VERSION : 0.1
   VAR_TEMP   // added for the SCL form of the ladder/FBD networks
      _w1 : Bool;
      _s5time1 : S5Time;
   END_VAR
BEGIN

REGION Network 1: Aviso 1 - Falla Conexión con sensor de Temperatura torres de Cavaleto
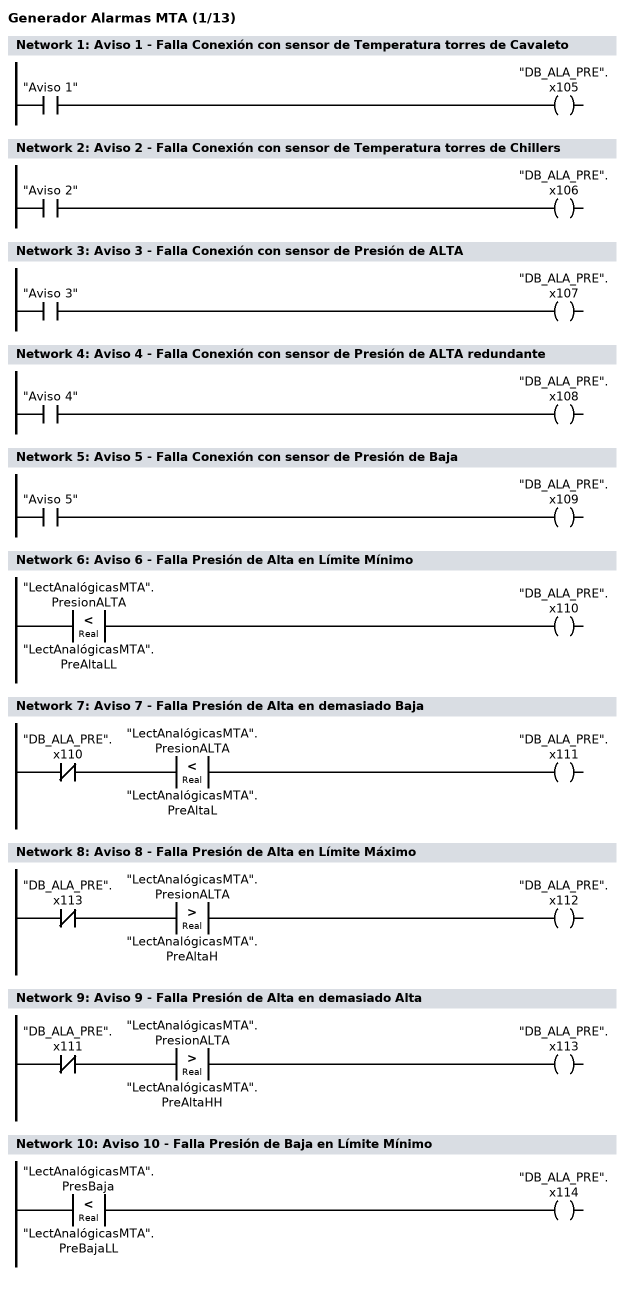
   RUNG wire#powerrail
      Contact( "Aviso 1" )
      Coil( "DB_ALA_PRE".x105 )
   END_RUNG
   // the same network as SCL:
   "DB_ALA_PRE".x105 := "Aviso 1";
END_REGION

REGION Network 2: Aviso 2 - Falla Conexión con sensor de Temperatura torres de Chillers
   RUNG wire#powerrail
      Contact( "Aviso 2" )
      Coil( "DB_ALA_PRE".x106 )
   END_RUNG
   // the same network as SCL:
   "DB_ALA_PRE".x106 := "Aviso 2";
END_REGION

REGION Network 3: Aviso 3 - Falla Conexión con sensor de Presión de ALTA
   RUNG wire#powerrail
      Contact( "Aviso 3" )
      Coil( "DB_ALA_PRE".x107 )
   END_RUNG
   // the same network as SCL:
   "DB_ALA_PRE".x107 := "Aviso 3";
END_REGION

REGION Network 4: Aviso 4 - Falla Conexión con sensor de Presión de ALTA redundante
   RUNG wire#powerrail
      Contact( "Aviso 4" )
      Coil( "DB_ALA_PRE".x108 )
   END_RUNG
   // the same network as SCL:
   "DB_ALA_PRE".x108 := "Aviso 4";
END_REGION

REGION Network 5: Aviso 5 - Falla Conexión con sensor de Presión de Baja
   RUNG wire#powerrail
      Contact( "Aviso 5" )
      Coil( "DB_ALA_PRE".x109 )
   END_RUNG
   // the same network as SCL:
   "DB_ALA_PRE".x109 := "Aviso 5";
END_REGION

REGION Network 6: Aviso 6 - Falla Presión de Alta en Límite Mínimo
   RUNG wire#powerrail
      { S7_Templates := "SrcType := Real" } LT_Contact(in1 := "LectAnalógicasMTA".PresionALTA, in2 := "LectAnalógicasMTA".PreAltaLL)
      Coil( "DB_ALA_PRE".x110 )
   END_RUNG
   // the same network as SCL:
   "DB_ALA_PRE".x110 := "LectAnalógicasMTA".PresionALTA < "LectAnalógicasMTA".PreAltaLL;
END_REGION

REGION Network 7: Aviso 7 - Falla Presión de Alta en demasiado Baja
   RUNG wire#powerrail
      I_Contact( "DB_ALA_PRE".x110 )
      { S7_Templates := "SrcType := Real" } LT_Contact(in1 := "LectAnalógicasMTA".PresionALTA, in2 := "LectAnalógicasMTA".PreAltaL)
      Coil( "DB_ALA_PRE".x111 )
   END_RUNG
   // the same network as SCL:
   "DB_ALA_PRE".x111 := NOT "DB_ALA_PRE".x110 AND ("LectAnalógicasMTA".PresionALTA < "LectAnalógicasMTA".PreAltaL);
END_REGION

REGION Network 8: Aviso 8 - Falla Presión de Alta en Límite Máximo
   RUNG wire#powerrail
      I_Contact( "DB_ALA_PRE".x113 )
      { S7_Templates := "SrcType := Real" } GT_Contact(in1 := "LectAnalógicasMTA".PresionALTA, in2 := "LectAnalógicasMTA".PreAltaH)
      Coil( "DB_ALA_PRE".x112 )
   END_RUNG
   // the same network as SCL:
   "DB_ALA_PRE".x112 := NOT "DB_ALA_PRE".x113 AND ("LectAnalógicasMTA".PresionALTA > "LectAnalógicasMTA".PreAltaH);
END_REGION

REGION Network 9: Aviso 9 - Falla Presión de Alta en demasiado Alta
   RUNG wire#powerrail
      I_Contact( "DB_ALA_PRE".x111 )
      { S7_Templates := "SrcType := Real" } GT_Contact(in1 := "LectAnalógicasMTA".PresionALTA, in2 := "LectAnalógicasMTA".PreAltaHH)
      Coil( "DB_ALA_PRE".x113 )
   END_RUNG
   // the same network as SCL:
   "DB_ALA_PRE".x113 := NOT "DB_ALA_PRE".x111 AND ("LectAnalógicasMTA".PresionALTA > "LectAnalógicasMTA".PreAltaHH);
END_REGION

REGION Network 10: Aviso 10 - Falla Presión de Baja en Límite Mínimo
   RUNG wire#powerrail
      { S7_Templates := "SrcType := Real" } LT_Contact(in1 := "LectAnalógicasMTA".PresBaja, in2 := "LectAnalógicasMTA".PreBajaLL)
      Coil( "DB_ALA_PRE".x114 )
   END_RUNG
   // the same network as SCL:
   "DB_ALA_PRE".x114 := "LectAnalógicasMTA".PresBaja < "LectAnalógicasMTA".PreBajaLL;
END_REGION

REGION Network 11: Aviso 11 - Falla Presión de Baja en demasiado Baja
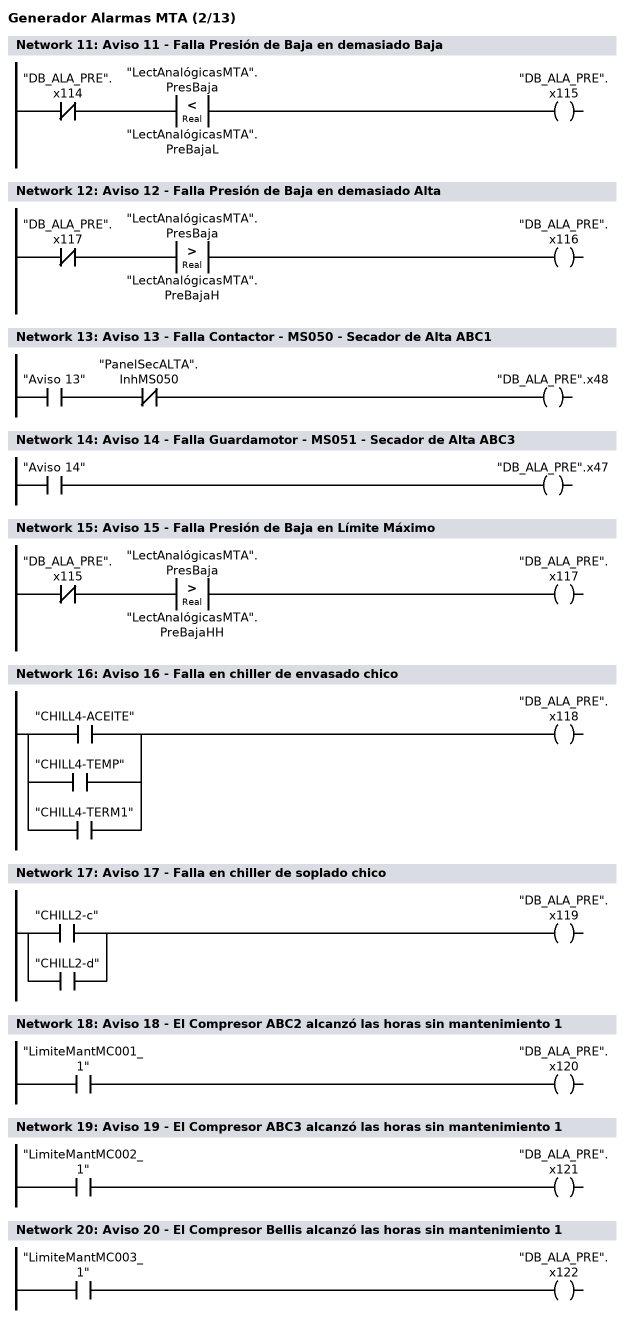
   RUNG wire#powerrail
      I_Contact( "DB_ALA_PRE".x114 )
      { S7_Templates := "SrcType := Real" } LT_Contact(in1 := "LectAnalógicasMTA".PresBaja, in2 := "LectAnalógicasMTA".PreBajaL)
      Coil( "DB_ALA_PRE".x115 )
   END_RUNG
   // the same network as SCL:
   "DB_ALA_PRE".x115 := NOT "DB_ALA_PRE".x114 AND ("LectAnalógicasMTA".PresBaja < "LectAnalógicasMTA".PreBajaL);
END_REGION

REGION Network 12: Aviso 12 - Falla Presión de Baja en demasiado Alta
   RUNG wire#powerrail
      I_Contact( "DB_ALA_PRE".x117 )
      { S7_Templates := "SrcType := Real" } GT_Contact(in1 := "LectAnalógicasMTA".PresBaja, in2 := "LectAnalógicasMTA".PreBajaH)
      Coil( "DB_ALA_PRE".x116 )
   END_RUNG
   // the same network as SCL:
   "DB_ALA_PRE".x116 := NOT "DB_ALA_PRE".x117 AND ("LectAnalógicasMTA".PresBaja > "LectAnalógicasMTA".PreBajaH);
END_REGION

REGION Network 13: Aviso 13 - Falla Contactor - MS050 - Secador de Alta ABC1
   RUNG wire#powerrail
      Contact( "Aviso 13" )
      I_Contact( "PanelSecALTA".InhMS050 )
      Coil( "DB_ALA_PRE".x48 )
   END_RUNG
   // the same network as SCL:
   "DB_ALA_PRE".x48 := "Aviso 13" AND NOT "PanelSecALTA".InhMS050;
END_REGION

REGION Network 14: Aviso 14 - Falla Guardamotor - MS051 - Secador de Alta ABC3
   RUNG wire#powerrail
      Contact( "Aviso 14" )
      Coil( "DB_ALA_PRE".x47 )
   END_RUNG
   // the same network as SCL:
   "DB_ALA_PRE".x47 := "Aviso 14";
END_REGION

REGION Network 15: Aviso 15 - Falla Presión de Baja en Límite Máximo
   RUNG wire#powerrail
      I_Contact( "DB_ALA_PRE".x115 )
      { S7_Templates := "SrcType := Real" } GT_Contact(in1 := "LectAnalógicasMTA".PresBaja, in2 := "LectAnalógicasMTA".PreBajaHH)
      Coil( "DB_ALA_PRE".x117 )
   END_RUNG
   // the same network as SCL:
   "DB_ALA_PRE".x117 := NOT "DB_ALA_PRE".x115 AND ("LectAnalógicasMTA".PresBaja > "LectAnalógicasMTA".PreBajaHH);
END_REGION

REGION Network 16: Aviso 16 - Falla en chiller de envasado chico
   RUNG wire#powerrail
      Contact( "CHILL4-ACEITE" )
      wire#w1
      Coil( "DB_ALA_PRE".x118 )
   END_RUNG
   RUNG wire#powerrail
      Contact( "CHILL4-TEMP" )
   END_RUNG wire#w1
   RUNG wire#powerrail
      Contact( "CHILL4-TERM1" )
   END_RUNG wire#w1
   // the same network as SCL:
   "DB_ALA_PRE".x118 := "CHILL4-ACEITE" OR "CHILL4-TEMP" OR "CHILL4-TERM1";
END_REGION

REGION Network 17: Aviso 17 - Falla en chiller de soplado chico
   RUNG wire#powerrail
      Contact( "CHILL2-c" )
      wire#w1
      Coil( "DB_ALA_PRE".x119 )
   END_RUNG
   RUNG wire#powerrail
      Contact( "CHILL2-d" )
   END_RUNG wire#w1
   // the same network as SCL:
   "DB_ALA_PRE".x119 := "CHILL2-c" OR "CHILL2-d";
END_REGION

REGION Network 18: Aviso 18 - El Compresor ABC2 alcanzó las horas sin mantenimiento 1
   RUNG wire#powerrail
      Contact( "LimiteMantMC001_1" )
      Coil( "DB_ALA_PRE".x120 )
   END_RUNG
   // the same network as SCL:
   "DB_ALA_PRE".x120 := "LimiteMantMC001_1";
END_REGION

REGION Network 19: Aviso 19 - El Compresor ABC3 alcanzó las horas sin mantenimiento 1
   RUNG wire#powerrail
      Contact( "LimiteMantMC002_1" )
      Coil( "DB_ALA_PRE".x121 )
   END_RUNG
   // the same network as SCL:
   "DB_ALA_PRE".x121 := "LimiteMantMC002_1";
END_REGION

REGION Network 20: Aviso 20 - El Compresor Bellis alcanzó las horas sin mantenimiento 1
   RUNG wire#powerrail
      Contact( "LimiteMantMC003_1" )
      Coil( "DB_ALA_PRE".x122 )
   END_RUNG
   // the same network as SCL:
   "DB_ALA_PRE".x122 := "LimiteMantMC003_1";
END_REGION

REGION Network 21: Aviso 21 - El Compresor ABC4 alcanzó las horas sin mantenimiento 1
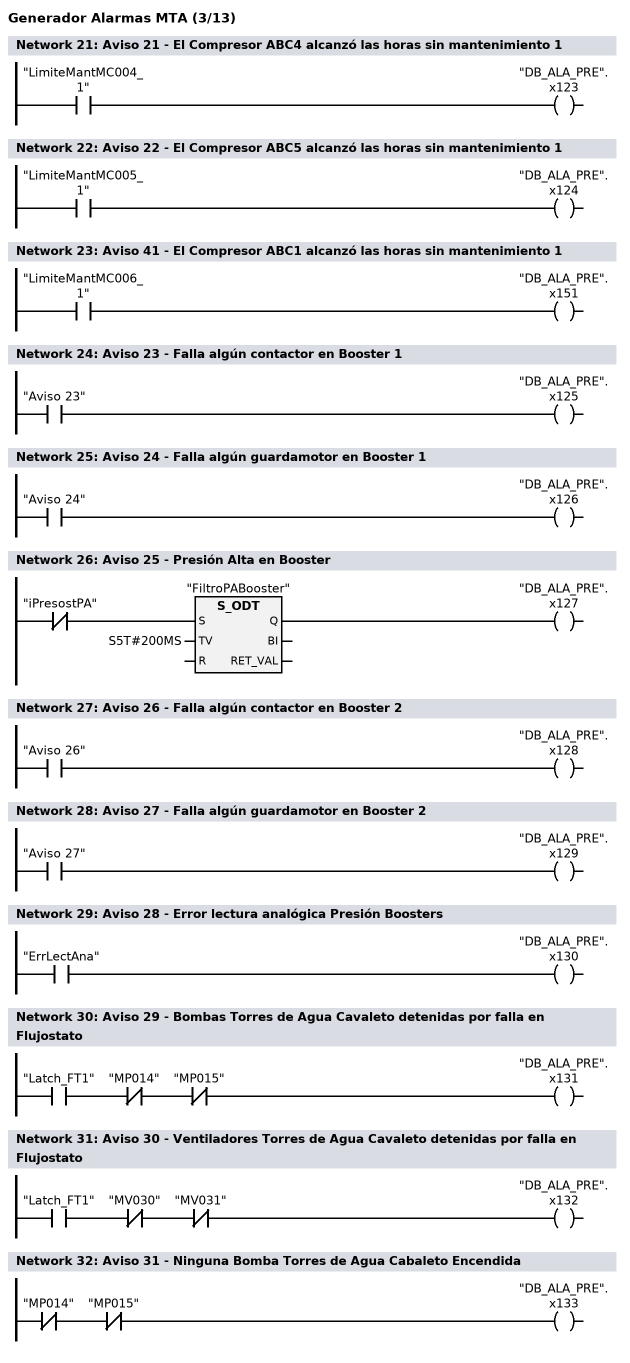
   RUNG wire#powerrail
      Contact( "LimiteMantMC004_1" )
      Coil( "DB_ALA_PRE".x123 )
   END_RUNG
   // the same network as SCL:
   "DB_ALA_PRE".x123 := "LimiteMantMC004_1";
END_REGION

REGION Network 22: Aviso 22 - El Compresor ABC5 alcanzó las horas sin mantenimiento 1
   RUNG wire#powerrail
      Contact( "LimiteMantMC005_1" )
      Coil( "DB_ALA_PRE".x124 )
   END_RUNG
   // the same network as SCL:
   "DB_ALA_PRE".x124 := "LimiteMantMC005_1";
END_REGION

REGION Network 23: Aviso 41 - El Compresor ABC1 alcanzó las horas sin mantenimiento 1
   RUNG wire#powerrail
      Contact( "LimiteMantMC006_1" )
      Coil( "DB_ALA_PRE".x151 )
   END_RUNG
   // the same network as SCL:
   "DB_ALA_PRE".x151 := "LimiteMantMC006_1";
END_REGION

REGION Network 24: Aviso 23 - Falla algún contactor en Booster 1
   RUNG wire#powerrail
      Contact( "Aviso 23" )
      Coil( "DB_ALA_PRE".x125 )
   END_RUNG
   // the same network as SCL:
   "DB_ALA_PRE".x125 := "Aviso 23";
END_REGION

REGION Network 25: Aviso 24 - Falla algún guardamotor en Booster 1
   RUNG wire#powerrail
      Contact( "Aviso 24" )
      Coil( "DB_ALA_PRE".x126 )
   END_RUNG
   // the same network as SCL:
   "DB_ALA_PRE".x126 := "Aviso 24";
END_REGION

REGION Network 26: Aviso 25 - Presión Alta en Booster
   RUNG wire#powerrail
      I_Contact( "iPresostPA" )
      S_ODT(T_NO := "FiltroPABooster", TV := S5T#200MS, R :=, BI =>, RET_VAL =>)
      Coil( "DB_ALA_PRE".x127 )
   END_RUNG
   // the same network as SCL:
   #_s5time1 := S_ODT(T_NO := "FiltroPABooster", S := NOT "iPresostPA", TV := S5T#200MS, Q => #_w1);
   "DB_ALA_PRE".x127 := #_w1;
END_REGION

REGION Network 27: Aviso 26 - Falla algún contactor en Booster 2
   RUNG wire#powerrail
      Contact( "Aviso 26" )
      Coil( "DB_ALA_PRE".x128 )
   END_RUNG
   // the same network as SCL:
   "DB_ALA_PRE".x128 := "Aviso 26";
END_REGION

REGION Network 28: Aviso 27 - Falla algún guardamotor en Booster 2
   RUNG wire#powerrail
      Contact( "Aviso 27" )
      Coil( "DB_ALA_PRE".x129 )
   END_RUNG
   // the same network as SCL:
   "DB_ALA_PRE".x129 := "Aviso 27";
END_REGION

REGION Network 29: Aviso 28 - Error lectura analógica Presión Boosters
   RUNG wire#powerrail
      Contact( "ErrLectAna" )
      Coil( "DB_ALA_PRE".x130 )
   END_RUNG
   // the same network as SCL:
   "DB_ALA_PRE".x130 := "ErrLectAna";
END_REGION

REGION Network 30: Aviso 29 - Bombas Torres de Agua Cavaleto detenidas por falla en Flujostato
   RUNG wire#powerrail
      Contact( "Latch_FT1" )
      I_Contact( "MP014" )
      I_Contact( "MP015" )
      Coil( "DB_ALA_PRE".x131 )
   END_RUNG
   // the same network as SCL:
   "DB_ALA_PRE".x131 := "Latch_FT1" AND NOT "MP014" AND NOT "MP015";
END_REGION

REGION Network 31: Aviso 30 - Ventiladores Torres de Agua Cavaleto detenidas por falla en Flujostato
   RUNG wire#powerrail
      Contact( "Latch_FT1" )
      I_Contact( "MV030" )
      I_Contact( "MV031" )
      Coil( "DB_ALA_PRE".x132 )
   END_RUNG
   // the same network as SCL:
   "DB_ALA_PRE".x132 := "Latch_FT1" AND NOT "MV030" AND NOT "MV031";
END_REGION

REGION Network 32: Aviso 31 - Ninguna Bomba Torres de Agua Cabaleto Encendida
   RUNG wire#powerrail
      I_Contact( "MP014" )
      I_Contact( "MP015" )
      Coil( "DB_ALA_PRE".x133 )
   END_RUNG
   // the same network as SCL:
   "DB_ALA_PRE".x133 := NOT "MP014" AND NOT "MP015";
END_REGION

REGION Network 33: Aviso 32 - Compresores Alta Detenidos por Flujostato Torres de Agua Cabaleto
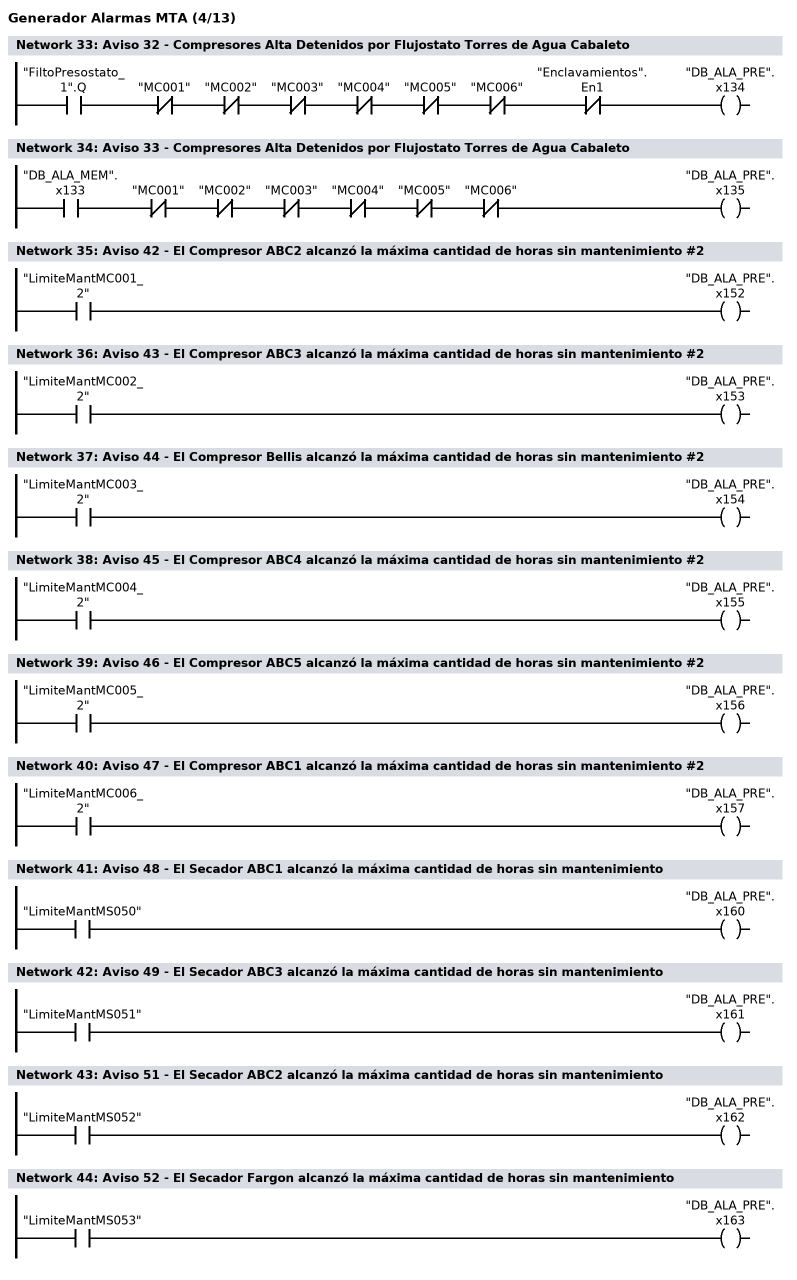
   RUNG wire#powerrail
      Contact( "FiltoPresostato_1".Q )
      I_Contact( "MC001" )
      I_Contact( "MC002" )
      I_Contact( "MC003" )
      I_Contact( "MC004" )
      I_Contact( "MC005" )
      I_Contact( "MC006" )
      I_Contact( "Enclavamientos".En1 )
      Coil( "DB_ALA_PRE".x134 )
   END_RUNG
   // the same network as SCL:
   "DB_ALA_PRE".x134 := "FiltoPresostato_1".Q AND NOT "MC001" AND NOT "MC002" AND NOT "MC003" AND NOT "MC004" AND NOT "MC005" AND NOT "MC006" AND NOT "Enclavamientos".En1;
END_REGION

REGION Network 34: Aviso 33 - Compresores Alta Detenidos por Flujostato Torres de Agua Cabaleto
   RUNG wire#powerrail
      Contact( "DB_ALA_MEM".x133 )
      I_Contact( "MC001" )
      I_Contact( "MC002" )
      I_Contact( "MC003" )
      I_Contact( "MC004" )
      I_Contact( "MC005" )
      I_Contact( "MC006" )
      Coil( "DB_ALA_PRE".x135 )
   END_RUNG
   // the same network as SCL:
   "DB_ALA_PRE".x135 := "DB_ALA_MEM".x133 AND NOT "MC001" AND NOT "MC002" AND NOT "MC003" AND NOT "MC004" AND NOT "MC005" AND NOT "MC006";
END_REGION

REGION Network 35: Aviso 42 - El Compresor ABC2 alcanzó la máxima cantidad de horas sin mantenimiento #2
   RUNG wire#powerrail
      Contact( "LimiteMantMC001_2" )
      Coil( "DB_ALA_PRE".x152 )
   END_RUNG
   // the same network as SCL:
   "DB_ALA_PRE".x152 := "LimiteMantMC001_2";
END_REGION

REGION Network 36: Aviso 43 - El Compresor ABC3 alcanzó la máxima cantidad de horas sin mantenimiento #2
   RUNG wire#powerrail
      Contact( "LimiteMantMC002_2" )
      Coil( "DB_ALA_PRE".x153 )
   END_RUNG
   // the same network as SCL:
   "DB_ALA_PRE".x153 := "LimiteMantMC002_2";
END_REGION

REGION Network 37: Aviso 44 - El Compresor Bellis alcanzó la máxima cantidad de horas sin mantenimiento #2
   RUNG wire#powerrail
      Contact( "LimiteMantMC003_2" )
      Coil( "DB_ALA_PRE".x154 )
   END_RUNG
   // the same network as SCL:
   "DB_ALA_PRE".x154 := "LimiteMantMC003_2";
END_REGION

REGION Network 38: Aviso 45 - El Compresor ABC4 alcanzó la máxima cantidad de horas sin mantenimiento #2
   RUNG wire#powerrail
      Contact( "LimiteMantMC004_2" )
      Coil( "DB_ALA_PRE".x155 )
   END_RUNG
   // the same network as SCL:
   "DB_ALA_PRE".x155 := "LimiteMantMC004_2";
END_REGION

REGION Network 39: Aviso 46 - El Compresor ABC5 alcanzó la máxima cantidad de horas sin mantenimiento #2
   RUNG wire#powerrail
      Contact( "LimiteMantMC005_2" )
      Coil( "DB_ALA_PRE".x156 )
   END_RUNG
   // the same network as SCL:
   "DB_ALA_PRE".x156 := "LimiteMantMC005_2";
END_REGION

REGION Network 40: Aviso 47 - El Compresor ABC1 alcanzó la máxima cantidad de horas sin mantenimiento #2
   RUNG wire#powerrail
      Contact( "LimiteMantMC006_2" )
      Coil( "DB_ALA_PRE".x157 )
   END_RUNG
   // the same network as SCL:
   "DB_ALA_PRE".x157 := "LimiteMantMC006_2";
END_REGION

REGION Network 41: Aviso 48 - El Secador ABC1 alcanzó la máxima cantidad de horas sin mantenimiento
   RUNG wire#powerrail
      Contact( "LimiteMantMS050" )
      Coil( "DB_ALA_PRE".x160 )
   END_RUNG
   // the same network as SCL:
   "DB_ALA_PRE".x160 := "LimiteMantMS050";
END_REGION

REGION Network 42: Aviso 49 - El Secador ABC3 alcanzó la máxima cantidad de horas sin mantenimiento
   RUNG wire#powerrail
      Contact( "LimiteMantMS051" )
      Coil( "DB_ALA_PRE".x161 )
   END_RUNG
   // the same network as SCL:
   "DB_ALA_PRE".x161 := "LimiteMantMS051";
END_REGION

REGION Network 43: Aviso 51 - El Secador ABC2 alcanzó la máxima cantidad de horas sin mantenimiento
   RUNG wire#powerrail
      Contact( "LimiteMantMS052" )
      Coil( "DB_ALA_PRE".x162 )
   END_RUNG
   // the same network as SCL:
   "DB_ALA_PRE".x162 := "LimiteMantMS052";
END_REGION

REGION Network 44: Aviso 52 - El Secador Fargon alcanzó la máxima cantidad de horas sin mantenimiento
   RUNG wire#powerrail
      Contact( "LimiteMantMS053" )
      Coil( "DB_ALA_PRE".x163 )
   END_RUNG
   // the same network as SCL:
   "DB_ALA_PRE".x163 := "LimiteMantMS053";
END_REGION

REGION Network 45: Aviso 54 - El Secador Sullair 1 alcanzó la máxima cantidad de horas sin mantenimiento 1
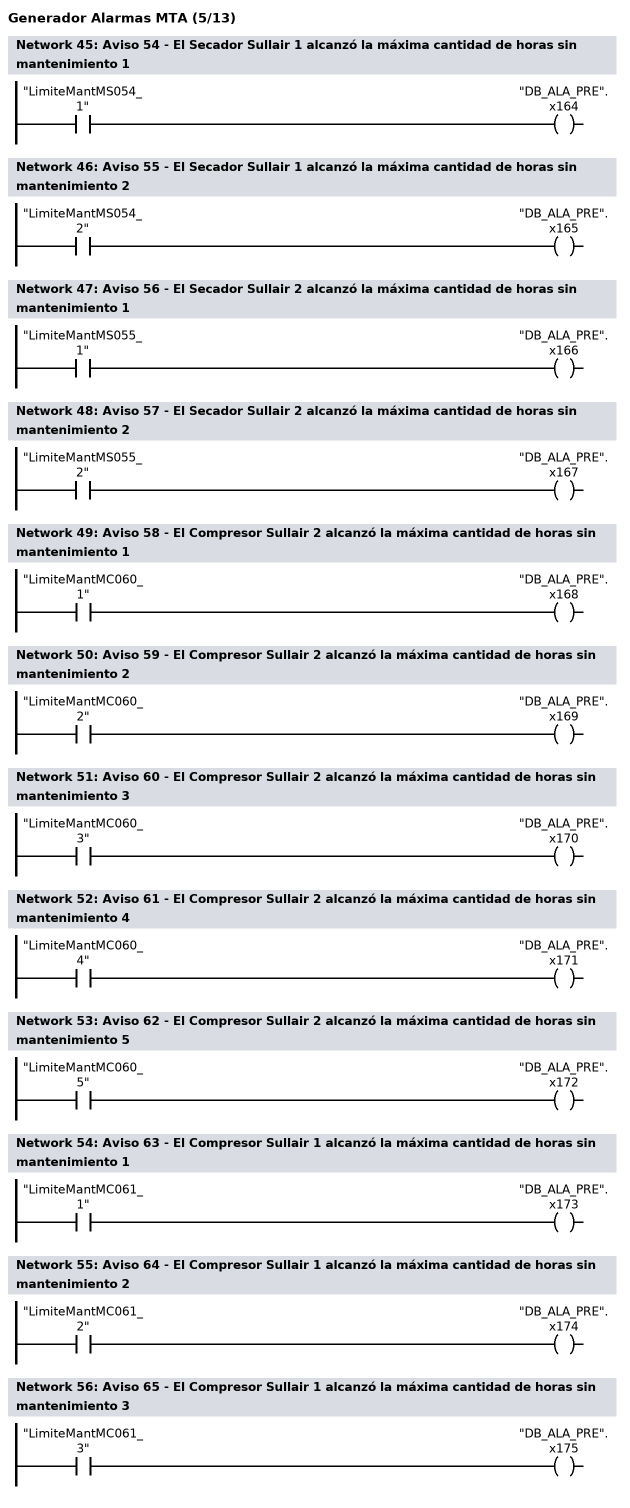
   RUNG wire#powerrail
      Contact( "LimiteMantMS054_1" )
      Coil( "DB_ALA_PRE".x164 )
   END_RUNG
   // the same network as SCL:
   "DB_ALA_PRE".x164 := "LimiteMantMS054_1";
END_REGION

